VAR_GLOBAL   (* controller tags *)
   ACTIVE_MODE : ALIAS FOR N54[208].3;
   AFI : ALIAS FOR B3[7].15;
   AFITC : ALIAS FOR B3[15].15;
   AMAX_LEHR_SPD : ALIAS FOR I[81];
   APC_HOST_PERM : ALIAS FOR B3[0].7;
   AUX_xInitialize : BOOL;
   Axies : MOTION_GROUP; {access Read Only}
   B106 : DINT[1];
   B151 : DINT[20] := ([0] := 2#1111_1111_1111_1111_1111_1111_1111_1111, [1] := 2#1111_1111_1111_1111_1111_1111_1111_1111, [2] := 2#0000_0000_0000_0000_1111_1111_1111_1111);
        [0]   // Cross-break Zone 1 Bit shift file * INSIDE LEHR *
   B152 : DINT[50];
        [0]   // Cross-break Zone 2 Bit shift file ** LEHR EXIT **
        [8].14   // Crossbreak Zone 3 Crossbreak Active NEW Start bit
        [11].14   // Crossbreak Zone 3 Crossbreak Active OLD Start bit
   B153 : DINT[20] := ([0] := 2#1111_1111_1111_1111_1111_1111_1111_1111, [1] := 2#1111_1111_1111_1111_1111_1111_1111_1111, [2] := 2#1111_1111_1111_1111_1111_1111_1111_1111, [3] := 2#0000_0000_0000_0000_1111_1111_1111_1111);
        [0]   // Cross-break Zone 3 Bit shift file ** WASHER **
   B154 : DINT[20];
        [0]   // Cross-break Zone 4 Bit shift file * IMAGE AUTO *
        [1]   // Crossbreak
        [8].0   // Cross-break Zone 4 Bit shift file **
        [8].11   // Cross-break Zone 4 Bit shift file **
   B155 : DINT[20] := ([0] := 2#1111_1111_1111_1111_1111_1111_1111_1111, [1] := 2#1111_1111_1111_1111_1111_1111_1111_1111, [2] := 2#1111_1111_1111_1111_1111_1111_1111_1111, [3] := 2#1111_1111_1111_1111_1111_1111_1111_1111, [4] := 2#1111_1111_1111_1111_1111_1111_1111_1111, [5] := 2#1111_1111_1111_1111_1111_1111_1111_1111, [6] := 2#1111_1111_1111_1111_1111_1111_1111_1111, [7] := 2#1111_1111_1111_1111_1111_1111_1111_1111, [8] := 2#0000_0000_0000_0000_1111_1111_1111_1111);
        [0]   // Cross-break Zone 5 Bit shift file ** MAN. INSP **
        [1]   // Cross-break Zone 5 Bit shift file ** MAN. INSP **
        [1].11   // Cross-break Zone 5 Bit shift file APC Roll #1
        [4]   // Cross-break Zone 5 Bit shift file ** MAN. INSP **
        [4].0   // Cross-break Zone 5 Bit shift file APC Roll #2
        [5]   // Cross-break Zone 5 Bit shift file ** MAN. INSP **
   B175 : DINT[1];
   B176 : DINT[1] := ([0] := 2#0000_0000_0000_0000_0000_1100_0000_0000);
   B180 : DINT[10] := ([0] := 2#0000_0000_0000_0000_0000_1111_1000_0000, [1] := 2#0000_0000_0000_0000_0000_0000_0100_0000, [2] := 2#0000_0000_0000_0000_0000_0000_1000_0000, [4] := 2#0000_0000_0000_0000_0001_0000_0000_0000, [5] := 2#0000_0000_0000_0000_0000_0000_0011_0000);
   B3 : DINT[102] := ([0] := 2#0000_0000_0000_0000_0001_1001_0100_0000, [2] := 2#0000_0000_0000_0000_0000_0000_0000_0110, [7] := 2#0000_0000_0000_0000_0000_0000_0000_0001, [8] := 2#0000_0000_0000_0000_1100_0000_0000_0001, [10] := 2#0000_0000_0000_0000_0100_0000_0010_0001);
        [0].0   // Valid Flaw Data to Process
        [0].1   // Reversed Scanner
        [0].2   // Gun Number is Odd
        [0].3   // Cap Data Request ONS
        [0].4   // Reject (Flaw) PB ONS
        [0].5   // Gun Test Requested
        [0].7   // APC MACHINE Permissive to Run from Host
        [0].9   // HOST TRACKING Permissive to Operate lucor MSM machine
        [0].11   // Bridge in Down Position
        [0].12   // Bridge in Up Position
        [0].13   // Auto Down After Cross-Brk
        [0].14   // one shot
        [1].0   // one shot
        [1].1   // MARKING BRIDGE In final decel during downward travel
        [1].2   // No. 1 Crusher Chip Blower Manual Permissive
        [1].3   // No. 1 Crusher Chip Blower Automatic Permissive
        [1].12   // Cullet System M47B Fwd Direction Selected
        [1].13   // Cullet System M47B Rev Direction Selected
        [1].14   // Cullet System M37B Fwd Direction Selected
        [1].15   // Cullet Sytem M37B Rev Direction Selected
        [2].0   // One Shot
        [2].1   // ONE SHOT
        [2].2   // SPONGE ROLL MANUALLY ON
        [3].0   // Reliance Drive System Fault Permissive
        [3].1   // Cullet System Fault Permissive
        [4].0   // CROSS BREAK Present At Sub-surface Cutters
        [5].0   // temp debug for 1 m sync pulse
        [5].1   // temp debug for 1 m sync pulse
        [5].2   // LEHR SPEED Debug One shot
        [6].0   // One Shot for Accumulation of 20 50mm Pulses
        [6].1   // One Shot to Resume Accumulation of 50mm Pulses
        [7].0   // Crossbreak Active In Zones 1 or 2 Enable Beacons and Horn Lehr wall
        [7].15   // Always False
        [8].0   // Crossbreak 1 (Lehr) Fault Count One Shot
        [8].14   // North Chilled Water Blower Is Not On
        [8].15   // South Chilled Water Blower Is Not On
        [10].0   // APC Crossbreak or Estop Acknowledge to Reset Roller #1
        [10].1   // APC Early Crossbreak Drip Valve Shutoff
        [10].2   // LEHR SPEED one shot!
        [10].3   // LEHR SPEED one shot!
        [10].4   // Reliance Drive & Cullet System Alarm Horn Relay (Capping Rm)
        [10].5   // APC Crossbreak or Estop Acknowledge to Reset Roller #2
        [10].10   // APC Supply Flow Is Low Alarm
        [10].14   // Tony's Washer Disable Toggle Bit
        [10].15   // Always False
        [15].15   // Always false Tony Bit
        [80].0   // CT Lehr Conv have all stoped
        [0].6   // OK to Run Lehr AUX Conveyors
   B49 : DINT[100];
   B52 : DINT[100] := ([0] := 2#0000_0000_0000_0000_0000_0000_0000_0001);
        [0].0   // All of CT DRIVES Enable
   B73 : DINT[1];
        [0].1   // Two inch Tracking pulse For Lehr Speed
        [0].2   // Two inch Tracking pulse For trim Speed
   BIN_1B_EAST : ALIAS FOR O[112].12;
   BLOWER_ON : ALIAS FOR O[67].13;
   BOOTH_LIGHTS : ALIAS FOR N46[4];
   BRDG_EOT_LS_HI : ALIAS FOR I[12].3;
   BRDG_SLO_LS_HI : ALIAS FOR I[12].0;
   BRDG_SLO_LS_LO : ALIAS FOR I[12].1;
   BRIDGE_DOWN : ALIAS FOR B3[0].11;
   BRIDGE_DRV_FLT : ALIAS FOR I[17].0;
   BRIDGE_FIN_DEC : ALIAS FOR B3[1].1;
   BRIDGE_LO_LAMP : ALIAS FOR O[22].3;
   BRIDGE_MAN_INSP : ALIAS FOR I[18].4;
   BRIDGE_UP : ALIAS FOR B3[0].12;
   BRSH1_DN_FLT : ALIAS FOR I[43].1;
   BRSH1_DN_FWD : ALIAS FOR O[45].1;
   BRSH1_DN_REV : ALIAS FOR O[45].9;
   BRSH1_DN_SS1 : ALIAS FOR O[46].1;
   BRSH1_DN_SS2 : ALIAS FOR O[46].9;
   BRSH1_UP_FLT : ALIAS FOR I[43].0;
   BRSH1_UP_FWD : ALIAS FOR O[45].0;
   BRSH1_UP_REV : ALIAS FOR O[45].8;
   BRSH1_UP_SS1 : ALIAS FOR O[46].0;
   BRSH1_UP_SS2 : ALIAS FOR O[46].8;
   BRSH2_DN_FLT : ALIAS FOR I[43].3;
   BRSH2_DN_FWD : ALIAS FOR O[45].3;
   BRSH2_DN_REV : ALIAS FOR O[45].11;
   BRSH2_DN_SS1 : ALIAS FOR O[46].3;
   BRSH2_DN_SS2 : ALIAS FOR O[46].11;
   BRSH2_UP_FLT : ALIAS FOR I[43].2;
   BRSH2_UP_FWD : ALIAS FOR O[45].2;
   BRSH2_UP_REV : ALIAS FOR O[45].10;
   BRSH2_UP_SS1 : ALIAS FOR O[46].2;
   BRSH2_UP_SS2 : ALIAS FOR O[46].10;
   BT181_000 : MESSAGE;
        MessageParameters(ServiceCode := 16#004c, LocalElement := N125[0], ...)
   BT181_001 : MESSAGE;
        MessageParameters(ServiceCode := 16#004c, LocalElement := N125[62], ...)
   BT181_002 : MESSAGE;
        MessageParameters(ServiceCode := 16#004c, LocalElement := N125[123], ...)
   BT181_003 : MESSAGE;
        MessageParameters(ServiceCode := 16#004c, LocalElement := N125[183], ...)
   BT181_004 : MESSAGE;
        MessageParameters(ServiceCode := 16#004b, LocalElement := N124[0], ...)
   BT181_005 : MESSAGE;
        MessageParameters(ServiceCode := 16#004b, LocalElement := N124[62], ...)
   BT181_006 : MESSAGE;
        MessageParameters(ServiceCode := 16#004b, LocalElement := N124[123], ...)
   BT181_007 : MESSAGE;
        MessageParameters(ServiceCode := 16#004b, LocalElement := N124[183], ...)
   BT181_008 : MESSAGE;
        MessageParameters(ServiceCode := 16#004b, LocalElement := N124[250], ...)
   BT181_009 : MESSAGE;
        MessageParameters(ServiceCode := 16#004c, LocalElement := N125[350], ...)
   BT181_010 : MESSAGE;
        MessageParameters(ServiceCode := 16#004b, LocalElement := N124[350], ...)
   BT181_011 : MESSAGE;
   BT181_012 : MESSAGE;
        MessageParameters(LocalElement := N15[60], ...)
   BT181_013 : MESSAGE;   // MB TO M2 BT of MMI Data To New CLX PLC
        MessageParameters(LocalElement := N7[180], ...)
   BT181_014 : MESSAGE;   // M2 TO MB BT of MMI Data from New CLX PLC
        MessageParameters(LocalElement := N7[160], ...)
   BT41_000 : MESSAGE;   // VHSC BTR
        .EN   // VHSC BTR Enabled
        MessageParameters(ServiceCode := 16#004b, LocalElement := N42[71], ...)
   BT41_001 : MESSAGE;   // VHSC BTW
        .EN   // VHSC BTW Enabled
        MessageParameters(ServiceCode := 16#004c, LocalElement := N42[1], ...)
   BT41_002 : MESSAGE;
        MessageParameters(LocalElement := N45[21], ...)
   BT41_003 : MESSAGE;
        MessageParameters(LocalElement := N45[1], ...)
   BT41_004 : MESSAGE;
   BT41_005 : MESSAGE;
   BT41_006 : MESSAGE;   // Block Transfer Read Control for Analog Input Card in Washer Panel
        MessageParameters(ServiceCode := 16#004b, LocalElement := N61[1], ...)
   BT41_007 : MESSAGE;   // Block Transfer Write Control for Analog Input Card in Washer Panel
        MessageParameters(ServiceCode := 16#004c, LocalElement := N61[51], ...)
   C183 : COUNTER[3] := ([0].PRE := 1, [0].CU := 1, [1].PRE := 7, [1].CU := 1, [2].PRE := 3, [2].CU := 1);
   C1_ACK : ALIAS FOR N54[260].14;
   C1_ACTIVE_LAMP : ALIAS FOR N54[260].0;
   C1_BEACON : ALIAS FOR O[27].6;
   C1_BEACON2 : ALIAS FOR O[47].10;
   C1_HORN : ALIAS FOR O[27].5;
   C1_NTH_IN_LMP : ALIAS FOR N54[260].10;
   C1_NTH_IN_PE : ALIAS FOR N54[260].6;
   C1_NTH_IN_SS : ALIAS FOR N54[260].2;
   C1_NTH_OUT_LMP : ALIAS FOR N54[260].9;
   C1_NTH_OUT_PE : ALIAS FOR N54[260].5;
   C1_NTH_OUT_SS : ALIAS FOR N54[260].1;
   C1_PNL_FLT : ALIAS FOR I[113].2;
   C1_STH_IN_LMP : ALIAS FOR N54[260].12;
   C1_STH_IN_PE : ALIAS FOR N54[260].8;
   C1_STH_IN_SS : ALIAS FOR N54[260].4;
   C1_STH_OUT_LMP : ALIAS FOR N54[260].11;
   C1_STH_OUT_PE : ALIAS FOR N54[260].7;
   C1_STH_OUT_SS : ALIAS FOR N54[260].3;
   C253 : COUNTER[100];
   C2_ACTIVE_LAMP : ALIAS FOR N54[261].0;
   C2_NTH_IN_LMP : ALIAS FOR N54[261].10;
   C2_NTH_IN_PE : ALIAS FOR N54[261].6;
   C2_NTH_IN_SS : ALIAS FOR N54[261].2;
   C2_NTH_OUT_LMP : ALIAS FOR N54[261].9;
   C2_NTH_OUT_PE : ALIAS FOR N54[261].5;
   C2_NTH_OUT_SS : ALIAS FOR N54[261].1;
   C2_PNL_FLT : ALIAS FOR I[113].3;
   C2_STH_IN_LMP : ALIAS FOR N54[261].12;
   C2_STH_IN_PE : ALIAS FOR N54[261].8;
   C2_STH_IN_SS : ALIAS FOR N54[261].4;
   C2_STH_OUT_LMP : ALIAS FOR N54[261].11;
   C2_STH_OUT_PE : ALIAS FOR N54[261].7;
   C2_STH_OUT_SS : ALIAS FOR N54[261].3;
   C3_ACTIVE_LAMP : ALIAS FOR N54[262].0;
   C3_NTH_IN_LMP : ALIAS FOR N54[262].10;
   C3_NTH_IN_PE : ALIAS FOR N54[262].6;
   C3_NTH_IN_SS : ALIAS FOR N54[262].2;
   C3_NTH_OUT_LMP : ALIAS FOR N54[262].9;
   C3_NTH_OUT_PE : ALIAS FOR N54[262].5;
   C3_NTH_OUT_SS : ALIAS FOR N54[262].1;
   C3_PNL_FLT : ALIAS FOR I[113].4;
   C3_STH_IN_LMP : ALIAS FOR N54[262].12;
   C3_STH_IN_PE : ALIAS FOR N54[262].8;
   C3_STH_IN_SS : ALIAS FOR N54[262].4;
   C3_STH_OUT_LMP : ALIAS FOR N54[262].11;
   C3_STH_OUT_PE : ALIAS FOR N54[262].7;
   C3_STH_OUT_SS : ALIAS FOR N54[262].3;
   C3_STP : ALIAS FOR O[35].10;
   C4_NTH_IN_PE : ALIAS FOR N54[263].6;
   C4_NTH_IN_SS : ALIAS FOR N54[263].2;
   C4_NTH_OUT_PE : ALIAS FOR N54[263].5;
   C4_NTH_OUT_SS : ALIAS FOR N54[263].1;
   C4_PNL_FLT : ALIAS FOR I[113].1;
   C4_STH_IN_PE : ALIAS FOR N54[263].8;
   C4_STH_OUT_PE : ALIAS FOR N54[263].7;
   C5 : COUNTER[100] := ([0].PRE := 200, [1].PRE := 2, [2].PRE := 52, [2].ACC := 29, [3].PRE := 30000, [3].ACC := 2, [4].PRE := 30000, [5].PRE := 30000, [6].PRE := 1000, [6].ACC := 423, [7].PRE := 30000, [8].PRE := 1000, [8].ACC := 112, [8].CU := 1, [10].PRE := 30000, [12].PRE := 30000, [13].PRE := 32767, [13].ACC := 1912, [14].ACC := 74, [14].DN := 1, [15].ACC := 54, [15].DN := 1, [16].ACC := 33, [16].DN := 1, [17].ACC := 27, [17].DN := 1, [20].PRE := 1000, [20].ACC := 1748, [20].DN := 1, [21].PRE := 1000, [21].ACC := 13747, [21].DN := 1, [21].OV := 1, [25].PRE := 1000, [25].ACC := 853, [26].PRE := 10000, [26].ACC := 3, [27].PRE := 10000, [27].ACC := 4, [27].CU := 1, [28].PRE := 10000, [28].ACC := 4, [28].CU := 1, [29].PRE := 10000, [29].ACC := 4, [29].CU := 1, [30].PRE := 10000, [30].ACC := 4, [30].CU := 1, [31].PRE := 10000, [31].ACC := 2145, [32].PRE := 10000, [32].ACC := 4, [32].CU := 1, [33].PRE := 10000, [34].PRE := 10000, [34].ACC := 4, [35].PRE := 10000, [35].ACC := 2786, [36].PRE := 10000,
        [36].ACC := 4, [37].PRE := 10000, [37].ACC := 2743, [38].PRE := 10000, [38].ACC := 4, [39].PRE := 10000, [39].ACC := 2790, [40].PRE := 10000, [40].ACC := 4, [41].PRE := 10000, [41].ACC := 2693, [42].PRE := 10000, [42].ACC := 4, [43].PRE := 10000, [43].ACC := 5802, [44].PRE := 10000, [44].ACC := 4, [45].PRE := 10000, [45].ACC := 11749, [45].DN := 1, [46].PRE := 10000, [46].ACC := 4, [46].DN := 1, [46].OV := 1, [47].PRE := 10000, [47].ACC := 478, [48].PRE := 10000, [48].ACC := 4, [49].PRE := 10000, [49].ACC := 6623, [50].PRE := 10000, [50].ACC := 4424, [51].PRE := 10000, [51].ACC := 734, [52].PRE := 10000, [52].ACC := 5426, [53].PRE := 10000, [53].ACC := 783, [54].PRE := 10000, [54].ACC := 3735, [55].PRE := 10000, [55].ACC := 733, [56].PRE := 10000, [56].ACC := 3661, [57].PRE := 10000, [57].ACC := 727, [58].PRE := 1000, [58].ACC := 251, [58].CU := 1, [70].PRE := 10000, [70].CU := 1, [71].PRE := 10000, [71].ACC := 4, [71].CU := 1, [72].PRE := 10000, [72].CU := 1, [73].PRE := 10000, [73].ACC := 4, [73].CU := 1, [74].PRE := 10000,
        [74].CU := 1, [75].PRE := 10000, [75].ACC := 4, [75].CU := 1, [76].PRE := 10000, [76].CU := 1, [77].PRE := 10000, [77].ACC := 4, [77].CU := 1, [78].PRE := 1000, [78].ACC := 607, [79].PRE := 1000, [79].ACC := 300, [80].PRE := 1000, [80].ACC := 337, [81].PRE := 1000, [81].ACC := 1033, [81].DN := 1, [82].PRE := 1000, [82].ACC := 146, [83].PRE := 1000, [83].ACC := 63, [84].PRE := 1000, [84].ACC := 2159, [84].DN := 1, [85].PRE := 1000, [85].ACC := 553, [90].PRE := 10000, [90].ACC := 8, [91].PRE := 10000, [93].PRE := 1000, [93].ACC := 338, [93].CU := 1, [94].PRE := 100, [95].PRE := 100, [96].PRE := 100, [96].ACC := 65, [97].PRE := 100, [97].ACC := 65, [98].PRE := 10000, [98].ACC := 6222, [99].PRE := 1000, [99].ACC := 520, [99].CU := 1);
        [6]   // TEMP Counter for Number of Times South OUT Sensor gets Disabled
        [13]   // Reliance Drive & Cullet System Alarm Horn (Capping) Conter
        [20]   // DEBUG: Number Of Times Capping Lehr Speed is Greater than Automax Speed plus 15IPM
        [21]   // TEMP DEBUG NUMBER OF TIMES 1M SYNC PULSE PERIOD IS LESS THAN 8 SEC
        [25]   // M2-->>MB Counts number of Times Mainline Backup to Trim Deck Occurs
        [26]   // CB Zone 1 (Lehr) North Outside Debounce Counter
        [27]   // CB Zone 1 (Lehr) North Outside Fault Counter
        [28]   // CB Zone 1 (Lehr) North Inside Debounce Counter
        [29]   // CB Zone 1 (Lehr) North Inside Fault Counter
        [30]   // CB Zone 1 (Lehr) South Outside Debounce Counter
        [31]   // CB Zone 1 (Lehr) South Outside Fault Counter
        [32]   // CB Zone 1 (Lehr) South Inside Debounce Counter
        [33]   // CB Zone 1 (Lehr) South Inside Fault Counter
        [34]   // CB Zone 2 (Crusher 1) North Outside Debounce Counter
        [35]   // CB Zone 2 (Crusher 1) North Outside Fault Counter
        [36]   // CB Zone 2 (Crusher 1) North Inside Debounce Counter
        [37]   // CB Zone 2 (Crusher 1) North Inside Fault Counter
        [38]   // CB Zone 2 (Crusher 1) South Outside Debounce Counter
        [39]   // CB Zone 2 (Crusher 1) South Outside Fault Counter
        [40]   // CB Zone 2 (Crusher 1) South Inside Debounce Counter
        [41]   // CB Zone 2 (Crusher 1) South Inside Fault Counter
        [42]   // CB Zone 3 (washer) North Outside Debounce Counter
        [43]   // CB Zone 3 (washer) North Outside Fault Counter
        [44]   // CB Zone 3 (washer) North Inside Debounce Counter
        [45]   // CB Zone 3 (washer) North Inside Fault Counter
        [45].ACC   // Z2 NO
        [46]   // CB Zone 3 (washer) South Outside Debounce Counter
        [46].ACC   // Z2 NI
        [47]   // CB Zone 3 (washer) South Outside Fault Counter
        [47].ACC   // Z2 SO
        [48]   // CB Zone 3 (washer) South Inside Debounce Counter
        [48].ACC   // Z2 SI
        [49]   // CB Zone 3 (washer) South Inside Fault Counter
        [50].ACC   // Z3 NO
        [51]   // CB Zone 4 (Inspection Booth) North Outside Fault Counter
        [51].ACC   // Z3 NI
        [52].ACC   // Z3 SO
        [53]   // CB Zone 4 (Inspection Booth) North Inside Fault Counter
        [53].ACC   // Z3 NI
        [54].ACC   // Z4 SI
        [55]   // CB Zone 4 (Inspection Booth) South Outside Fault Counter
        [55].ACC   // Z4 SO
        [56].ACC   // Z4 NI
        [57]   // CB Zone 4 (Inspection Booth) South Inside Fault Counter
        [57].ACC   // Z4 NO
        [71].ACC   // Z5 NO
        [73].ACC   // Z5 SI
        [75].ACC   // Z5 SO
        [77].ACC   // Z5 SI
        [90]   // Temporary Counter to Monitor CT Master Drive Fault Contact 0 ON 03/11/08
        [94]   // I/O STATUS FILE: Rack 12 Group 6 FAULT
        [95]   // I/O STATUS FILE: Rack 12 Group 4 FAULT
        [96]   // I/O STATUS FILE: Rack 12 Group 2 FAULT
        [97]   // I/O STATUS FILE: Rack 12 Group 0 FAULT
        [98]   // Glass Travel Pulse Count (Counts 50mm Pulses reset @ 10000)
        [99]   // BRUSH 1 DRIVE FAULTS
   C5_ACTIVE_LAMP : ALIAS FOR N54[264].0;
   C5_MARKING_CB : ALIAS FOR N54[264].15;
   C5_NTH_IN_LMP : ALIAS FOR N54[264].10;
   C5_NTH_IN_PE : ALIAS FOR N54[264].6;
   C5_NTH_IN_SS : ALIAS FOR N54[264].2;
   C5_NTH_OUT_LMP : ALIAS FOR N54[264].9;
   C5_NTH_OUT_PE : ALIAS FOR N54[264].5;
   C5_NTH_OUT_SS : ALIAS FOR N54[264].1;
   C5_STH_IN_LMP : ALIAS FOR N54[264].12;
   C5_STH_IN_PE : ALIAS FOR N54[264].8;
   C5_STH_IN_SS : ALIAS FOR N54[264].4;
   C5_STH_OUT_LMP : ALIAS FOR N54[264].11;
   C5_STH_OUT_PE : ALIAS FOR N54[264].7;
   C5_STH_OUT_SS : ALIAS FOR N54[264].3;
   CAP_AHR_TMR : ALIAS FOR T4[6];
   CAP_ALM_HORN : ALIAS FOR O[11].2;
   CAW_OK_BIT_W_PLC : ALIAS FOR N251[901].0;
   CAWSV_ON_BIT_TO_WPLC : ALIAS FOR N251[900].0;
   CB_AT_SS_CUTTERS : ALIAS FOR B3[4].0;
   CBF_START_B : ALIAS FOR I[65].5;
   CBF_START_T : ALIAS FOR I[65].4;
   CBF_STOP_B : ALIAS FOR I[65].7;
   CBF_STOP_T : ALIAS FOR I[65].6;
   CHIP_BLOW_A : ALIAS FOR B3[1].3;
   CHIP_BLOW_M : ALIAS FOR B3[1].2;
   CHIP_BLOW_TMR : ALIAS FOR T51[9];
   CNV10_PROCST : ALIAS FOR I[19].9;
   CNV11_PROCST : ALIAS FOR I[3].1;
   CNV12_PROCST : ALIAS FOR I[3].2;
   CNV13_PROCST : ALIAS FOR I[3].3;
   CNV14_PROCST : ALIAS FOR I[3].4;
   CNV15_PROCST : ALIAS FOR I[3].5;
   CNV16_PROCST : ALIAS FOR I[3].7;
   CNV17_PROCST : ALIAS FOR I[3].8;
   CNV1_PROCST : ALIAS FOR I[19].0;
   CNV2_PROCST : ALIAS FOR I[19].1;
   CNV3_PROCST : ALIAS FOR I[19].2;
   CNV4_PROCST : ALIAS FOR I[19].3;
   CNV5_PROCST : ALIAS FOR I[19].4;
   CNV6_PROCST : ALIAS FOR I[19].5;
   CNV7_PROCST : ALIAS FOR I[19].6;
   CNV8_PROCST : ALIAS FOR I[19].7;
   CNV9_PROCST : ALIAS FOR I[19].8;
   ConsumedFromCullet : UDT_CONSUMED_CULLET;
   ConsumedFromMCC1300 : UDT_CONSUMED_NEXT := (iM2toMB_2 := 132, iM2toMB_4 := 2048);
   CPU_FaultRecord : SYS_FaultRecord;
   CPU_LastFaultRecord : SYS_FaultRecord;
   CR1_0FF_LAMP : ALIAS FOR O[67].9;
   CR1_ALM : ALIAS FOR I[65].1;
   CR1_AUTO : ALIAS FOR I[64].13;
   CR1_AUTO_MODE : ALIAS FOR N54[240].1;
   CR1_CONT_FAIL : ALIAS FOR N54[240].4;
   CR1_CULLET_FAIL : ALIAS FOR N54[240].6;
   CR1_DNET_SS1 : ALIAS FOR N179[18];
   CR1_DNET_SS2 : ALIAS FOR N179[30];
   CR1_DOWN_PROX : ALIAS FOR I[64].11;
   CR1_DOWN_PWRLOS : ALIAS FOR N54[240].10;
   CR1_DOWN_RLY : ALIAS FOR O[67].1;
   CR1_DROP_COND : ALIAS FOR N54[240].13;
   CR1_DRV_FLT_LMP : ALIAS FOR O[66].8;
   CR1_DRV_FLT_RLY : ALIAS FOR O[66].9;
   CR1_DWN_PROX : ALIAS FOR N54[240].14;
   CR1_ESTOP : ALIAS FOR N54[240].3;
   CR1_FLT : ALIAS FOR I[65].0;
   CR1_FRSTSCN_TMR : ALIAS FOR T51[11];
   CR1_FWD : ALIAS FOR O[66].0;
   CR1_MAN_LOWER : ALIAS FOR I[64].15;
   CR1_MAN_MODE : ALIAS FOR N54[240].2;
   CR1_MAN_RAISE : ALIAS FOR I[64].14;
   CR1_NODROP_COND : ALIAS FOR N54[240].0;
   CR1_ON_LAMP : ALIAS FOR O[67].8;
   CR1_RUN_ENABLE : ALIAS FOR O[117].4;
   CR1_SS1 : ALIAS FOR O[66].2;
   CR1_SS2 : ALIAS FOR O[66].4;
   CR1_SS3 : ALIAS FOR O[66].6;
   CR1_START_PB : ALIAS FOR I[65].12;
   CR1_STOP_PB : ALIAS FOR I[65].13;
   CR1_TEST_PB : ALIAS FOR I[65].3;
   CR1_UP_PROX : ALIAS FOR I[64].12;
   CR1_UP_RLY : ALIAS FOR O[67].0;
   CR1_UPT_PROX : ALIAS FOR N54[240].15;
   CULL_FLT : ALIAS FOR B3[3].1;
   CULLET_FLT_PL : ALIAS FOR O[11].1;
   CURR_LSD : ALIAS FOR N42[74];
   CURR_MSD : ALIAS FOR N42[73];
   CURR_SYNC : ALIAS FOR N7[2];
   DateTime : DINT[7] := ([0] := 2023, [1] := 6, [2] := 9, [3] := 15, [4] := 17, [5] := 5, [6] := 737882);   // DINT array tag for retrieve wallclock time through GSV created during conversion
        [0]   // Year
        [1]   // Month
        [2]   // Day
        [3]   // Hour
        [4]   // Minute
        [5]   // Second
        [6]   // Microsecond
   DISABLE_REL : ALIAS FOR N46[3];
   DISTANCE : ALIAS FOR N7[1];
   DIV_POSITION : ALIAS FOR I[24].12;
   DIVERTER_POS1 : ALIAS FOR O[116].8;
   DRIVE_FAULT_PRESENT : BOOL; {access Read Only}
   ECLIPSE_OFF : ALIAS FOR N54[208].2;
   ECLIPSE_ON : ALIAS FOR N54[208].1;
   EMERGENCY_OK : BOOL;
   F58 : REAL[20] := ([0] := 5063.717);
        [0]   // APC Calculated Freq for APC Roller [Hz * 100]
   F74 : REAL[2] := ([0] := 13.333333, [1] := 0.15);
   F8 : REAL[20] := ([5] := 3.125);
        [5]   // SHEET TEMPERATURE: Tuning Factor to adjust PLC Value to match LED Display Unit
   F96 : REAL[50] := ([0] := 268.34647, [1] := 268.34647, [5] := 118.346466, [6] := 418.34647, [9] := 270.6, [10] := 270.6, [11] := 268.34647, [12] := 1.94725, [14] := 285.6, [20] := 268.34647, [21] := 268.34647, [22] := 268.34647, [23] := 268.34647, [24] := 268.34647, [25] := 268.34647, [26] := 268.34647, [27] := 268.34647, [28] := 268.34647, [29] := 268.34647, [30] := 270.6, [40] := 268.34647, [41] := 268.34647, [42] := 268.34647, [43] := 268.34647, [44] := 268.34647, [45] := 268.34647, [46] := 268.34647, [47] := 268.34647, [48] := 268.34647, [49] := 268.34647);
        [0]   // LEHR SPEED Current lehr Speed used Setting Speed of drives
        [1]   // LEHR SPEED Average lehr Speed Calculated from Sample table
        [5]   // LEHR SPEED Current Lehr Lower Limit
        [6]   // LEHR SPEED Current Lehr Speed upper Limit
        [9]   // LEHR SPEED Last lehr Speed Reset value
        [10]   // LEHR SPEED Information Received from Reliance AutoMax
        [11]   // LEHR SPEED Information Received from Reliance Capping system
        [14]   // DEBUG USAGE Lehr Speed from Automax Plus 15 IPM
        [20]   // LEHR SPEED Table of Speed samples Over last ten Seconds
        [21]   // LEHR SPEED Table of Lehr speed Samples over Ten seconds
   FAST_FLASH : ALIAS FOR T51[2];
   FFLASH_SLAVE : ALIAS FOR T51[3];
   FIRST_SCAN : ALIAS FOR S[1].15;
   FLAW_HEAD : ALIAS FOR N43[200];
   FLAW_LANE : ALIAS FOR N43[201];
   FLAW_OFF : ALIAS FOR N43[202];
   FLAW_OUT : ALIAS FOR N7[5];
   FLAW_POS : ALIAS FOR N7[4];
   FLAW_QUEUE : ALIAS FOR N7[9];
   FLAW_XLAT : ALIAS FOR N7[6];
   FLOW_CLK_LSD : ALIAS FOR N7[10];
   FLOW_CLK_MSD : ALIAS FOR N7[11];
   ForceStatus : INT;   // INT tag to retrieve Force enabled value through GSV created during conversion
   From_Cullet : DINT[10];
   GENERATOR_ON : ALIAS FOR N54[240].11;
   GENERATOR_RUN : ALIAS FOR I[65].15;
   GOOD_FLAW : ALIAS FOR B3[0].0;
   GP_M225_AccessArea : GP_AccessArea := (IN_xConditionOkAccess := 1); {access None}
   GP_M225_AccessArea_STC : GP_AccessArea_STC := (OSR_xRemoveAccess := 1, OSR_xRemoveAccessNotAccepted := 1, tmON_ForceAccess.PRE := 5000); {access None}
   GP_NetDiag : GP_NetworkDiag;
   GP_OB_InitializeDiag : GP_OB_Initialize := (OUT_dExecutionTime_ms := 500, OUT_dMaxExecutionTime_ms := 1033885, OUT_xOs_100ms := 1, OUT_xOs_200ms := 1, OUT_xOs_400ms := 1, OUT_xOs_500ms := 1, OUT_xOs_800ms := 1, OUT_xClock_100ms := 1, OUT_xClock_200ms := 1, OUT_xClock_400ms := 1, OUT_xClock_500ms := 1, OUT_xClock_800ms := 1, OUT_xClock_1s := 1, OUT_xClock_5s := 1, OUT_xClock_10s := 1, OUT_xClock_30s := 1, OUT_xClock_1h := 1, OUT_xDebugON := 1);
   GP_OB_InitializeDiag_STC : GP_OB_Initialize_STC := (dElapsed_1h_ms := 7496626, dElapsed_1min_ms := 56626, dElapsed_1s_ms := 626, dElapsed_2min_ms := 56626, dElapsed_2s_ms := 626, dElapsed_5s_ms := 1626, dElapsed_10min_ms := 296626, dElapsed_10s_ms := 6626, dElapsed_30min_ms := 296626, dElapsed_30s_ms := 26626, dElapsed_100ms_ms := 75523026, dElapsed_200ms_ms := 57149426, dElapsed_400ms_ms := 20402226, dElapsed_500ms_ms := 2028626, dElapsed_800ms_ms := 626, dlLastExecValue_us := 499964, rReminder_ms := -0.35214233, lwOldStartTime[0] := -592654905, lwOldStartTime[1] := 392627, lwStartTime[0] := -592654905, lwStartTime[1] := 392627);
   GP_OB_InitializeMain : GP_OB_Initialize := (OUT_dExecutionTime_ms := 10, OUT_dMaxExecutionTime_ms := 11, OUT_xOs_100ms := 1, OUT_xOs_200ms := 1, OUT_xClock_200ms := 1, OUT_xClock_800ms := 1, OUT_xClock_1s := 1, OUT_xClock_2s := 1, OUT_xClock_5s := 1, OUT_xClock_10s := 1, OUT_xClock_30s := 1, OUT_xClock_2min := 1, OUT_xClock_10min := 1, OUT_xDebugON := 1);
   GP_OB_InitializeMain_STC : GP_OB_Initialize_STC := (dElapsed_1h_ms := 4478668, dElapsed_1min_ms := 38668, dElapsed_1s_ms := 668, dElapsed_2min_ms := 38668, dElapsed_2s_ms := 668, dElapsed_5s_ms := 3668, dElapsed_10min_ms := 278668, dElapsed_10s_ms := 8668, dElapsed_30min_ms := 878668, dElapsed_30s_ms := 8668, dElapsed_100ms_ms := 68, dElapsed_200ms_ms := 68, dElapsed_400ms_ms := 268, dElapsed_500ms_ms := 168, dElapsed_800ms_ms := 268, dlLastExecValue_us := 9789, rReminder_ms := -0.0073947906, lwOldStartTime[0] := -593976054, lwOldStartTime[1] := 392627, lwStartTime[0] := -593976054, lwStartTime[1] := 392627);
   GUN_INDEX : ALIAS FOR N7[0];
   HMI_Alarm_Presence : BOOL;   // HMI_Alarm_Presence
   HMI_Alarm_Reset : BOOL;   // HMI_Alarm_Reset
   HMI_Alarms_0 : BOOL[32];   // HMI Alarms
   HMI_Alarms_1 : BOOL[32];   // HMI Alarms
   HMI_Alarms_2 : BOOL[32];   // HMI Alarms
   HMI_Alarms_3 : BOOL[32];   // HMI Alarms
   HMI_Alarms_4 : BOOL[32];   // HMI Alarms
   HMI_Alarms_5 : BOOL[32];   // HMI Alarms
   HMI_Alarms_6 : BOOL[32];   // HMI Alarms
   HMI_Alarms_7 : BOOL[32];   // HMI Alarms
   HMI_Alarms_8 : BOOL[32];   // HMI Alarms
   HMI_Alarms_9 : BOOL[32];   // HMI Alarms
   HMI_Always_ON : BOOL := 1;   // HMI Always ON
   HMI_MAN_CMD_WR : UDT_MAN_CMD_WR; {access Read Only}
   HMI_MOTOR_HMR : UDT_MOTOR_HMR; {access Read Only}
   HOST_DATA_REQ : ALIAS FOR N43[209].0;
   HOST_IAL_ALARM : ALIAS FOR N43[209].6;
   HOST_IAL_WD : ALIAS FOR N43[209].7;
   HOST_NWDATA_TMR : ALIAS FOR T4[3];
   I : INT[128] := ([14] := 2#0000_0000_0010_0001, [15] := 2#0000_0000_0010_0001, [16] := 2#0000_0000_0000_0100, [17] := 2#1001_0000_0100_0000, [42] := 2#0000_0100_1110_1110, [43] := 2#0000_0000_1011_0000, [49] := 2#0000_0000_0010_0001, [65] := 2#1000_0001_1100_0001, [80] := 2#0011_0110_1111_0011, [81] := 2#0000_1010_1001_0010, [83] := 2#0000_0000_0001_1111, [121] := 2#0000_0000_1000_0100, [123] := 2#0000_1000_0000_0000);
        [42].9   // VMCC W1 Alarm Reset (NOT USED ANYMORE)
        [62].14   // SPARE
        [120]   // M2 --> MB
        [0].15   // PANEL C1 M47B Conv Forward Selector (INCLINE)
        [1].8   // PANEL C1 M47B Conv Reverse Selector (INCLINE)
        [3].0   // Transfer 1 Belt Process Stop Enabled
        [3].1   // Conveyor 11 Process Stop Enabled
        [3].2   // Conveyor 12 Process Stop Enabled
        [3].3   // Conveyor 13 Process Stop Enabled
        [3].4   // Conveyor 14 Process Stop Enabled
        [3].5   // Conveyor 15 Process Stop Enabled
        [3].6   // Transfer 1A Bel Process Stop Enabled
        [3].7   // Conveyor 16 Process Stop Enabled
        [3].8   // Conveyor 17 Process Stop Enabled
        [12].0   // Bridge Top Slow Down L.S.
        [12].1   // Bridge bottom Slow L.S.
        [12].3   // Bridge Top E.O.T. L.S.
        [12].14   // Reliance Data Request
        [12].15   // Reliance Two inch Lehr Pulse
        [16].0   // ISRA 5D 24VDC OK
        [16].4   // ISRA 5D 12V DC OK
        [16].5   // ISRA 5D System Ok
        [16].6   // ISRA 5D System Warning
        [16].7   // ISRA 5D System Error 1
        [16].8   // ISRA 5D System Error 2
        [16].9   // VMCC MB Alarm Silence
        [16].10   // VMCC MB Alarm Reset
        [16].14   // ISRA 5D System Crossbreak
        [17].1   // South Chilled Water Blower Off PB I02105
        [17].2   // North Subsurface Cutter Alarm Signal
        [17].3   // South Subsurface Cutter Alarm Signal
        [17].4   // South Chilled Water Blower On PB I02104
        [17].5   // South Chilled Water Blower Off PB I02105
        [17].7   // South Chilled Water Blower VFD is Running Without Faults
        [17].9   // Inspection in Manual Mode
        [17].10   // North Chilled Water Blower On PB I02112
        [17].11   // North Chilled Water Blower Off PB I02113
        [16].3   // ISRA 5D System Watchdog (NOT USED)
        [17].13   // North Chilled Water Blower VFD is Running Without Faults
        [17].14   // TO BE VALORIZED FROM MCC1200 Data Request From New Cutting System (Data Request from Reliance)
        [18].2   // SPARE (APC Reset Button After Crossbreak)
        [18].4   // SPARE (Inspection in Manual Mode)
        [16].1   // Spare
        [18].3   // SPARE (APC ON/OFF (0=OFF) (1=ON))
        [19].0   // Conveyor 1 Process Stop Enabled
        [19].1   // Conveyor 2 Process Stop Enabled
        [19].2   // Conveyor 3 Process Stop Enabled
        [19].3   // Conveyor 4 Process Stop Enabled
        [19].4   // Conveyor 5 Process Stop Enabled
        [19].5   // Conveyor 6 Process Stop Enabled
        [19].6   // Conveyor 7 Process Stop Enabled
        [19].7   // Conveyor 8 Process Stop Enabled
        [19].8   // Conveyor 9 Process Stop Enabled
        [19].9   // Conveyor 10 Process Stop Enabled
        [24].0   // CRSSBRK ZONE 1 North Outside Bypass Switch
        [24].1   // CRSSBRK ZONE 1 North Inside Bypass Switch
        [24].2   // CRSSBRK ZONE 1 South Outside Bypass Switch
        [24].3   // CRSSBRK ZONE 1 South Inside Bypass Switch
        [24].4   // CRSSBRK ZONE 1 North Outside Photo-cell
        [24].5   // CRSSBRK ZONE 1 North Inside Photo-cell
        [24].6   // CRSSBRK ZONE 1 South Outside Photo-cell
        [24].7   // CRSSBRK ZONE 1 South Inside Photo-cell
        [24].8   // Cullet System M37B Fwd Direction Selector (Outside)
        [24].9   // Cullet System M37B Rev Direction Selector (Outside)
        [24].10   // Cullet System M47B Fwd Direction Selector (Outside)
        [24].11   // Cullet System M47B Rev Direction Selector (Outside)
        [24].12   // Diverter Position Selector At Cullet Op Panel
        [26].0   // CRSSBRK ZONE 2 North Outside Bypass Switch
        [26].1   // CRSSBRK ZONE 2 North Inside Bypass Switch
        [26].2   // CRSSBRK ZONE 2 South Outside Bypass Switch
        [26].3   // CRSSBRK ZONE 2 South Inside Bypass Switch
        [26].4   // CRSSBRK ZONE 2 North Outside Photo-cell
        [26].5   // CRSSBRK ZONE 2 North Inside Photo-cell
        [26].6   // CRSSBRK ZONE 2 South Outside Photo-cell
        [26].7   // CRSSBRK ZONE 2 South Inside Photo-cell
        [28].0   // CRSSBRK ZONE 3 North Outside Bypass Switch
        [28].1   // CRSSBRK ZONE 3 North Inside Bypass Switch
        [28].2   // CRSSBRK ZONE 3 South Outside Bypass Switch
        [28].3   // CRSSBRK ZONE 3 South Inside Bypass Switch
        [28].4   // CRSSBRK ZONE 3 North Outside Photo-cell
        [28].5   // CRSSBRK ZONE 3 North Inside Photo-cell
        [28].6   // CRSSBRK ZONE 3 South Outside Photo-cell
        [28].7   // CRSSBRK ZONE 3 South Inside Photo-cell
        [30].13   // CRSSBRK ZONE 4 Adapter power ON
        [30].15   // CRSSBRK ZONE 4 Output power ON
        [30].12   // IMAGE AUTO Retro-cover Closed Prox
        [32].0   // CRSSBRK ZONE 5 North Outside Bypass Switch
        [32].1   // CRSSBRK ZONE 5 North Inside Bypass Switch
        [32].2   // CRSSBRK ZONE 5 South Outside Bypass Switch
        [32].3   // CRSSBRK ZONE 5 South Inside Bypass Switch
        [32].4   // CRSSBRK ZONE 5 North Outside Photo-cell
        [32].5   // CRSSBRK ZONE 5 North Inside Photo-cell
        [32].6   // CRSSBRK ZONE 5 South Outside Photo-cell
        [32].7   // CRSSBRK ZONE 5 South Inside Photo-cell
        [32].8   // APC #1 Reset Button After Crossbreak
        [32].9   // APC Spray system OFF (1=OFF) (0=ON)
        [32].10   // APC #2 Reset Button After Crossbreak changed 22Mar2019TC
        [32].11   // APC Spray System Supply Flow Low (From SMC flow meter)
        [34].0   // MANUAL INSPCTN Booth Flaw Push-Button
        [34].1   // MANUAL INSPCTN Booth Reject Push-Button
        [34].3   // LOW-E Inspection Catwalk: Spray Zone 1 Pushbutton
        [34].4   // LOW-E Inspection Catwalk: Spray Zone 2 Pushbutton
        [34].5   // LOW-E Inspection Catwalk: Spray Zone 3 Pushbutton
        [34].6   // LOW-E Inspection Catwalk: Spray Zone 4 Pushbutton
        [34].7   // LOW-E Inspection Catwalk: Spray Zone 5 Pushbutton
        [34].8   // LOW-E Inspection Catwalk: Pulse Entire Ribbon Pushbutton
        [58].12   // SPARE
        [58].13   // SPARE
        [58].10   // SPARE
        [58].15   // SPARE
        [60].15   // SPARE
        [58].9   // SPARE
        [56].15   // SPARE
        [58].11   // SPARE
        [58].14   // SPARE
        [43].0   // VMCC W1 Upper Brush #1 Drive fault
        [43].1   // VMCC W1 Lower Brush #1 Drive fault
        [43].2   // VMCC W1 Upper Brush #2 Drive fault
        [43].3   // VMCC W1 Lower Brush #2 Drive fault
        [43].6   // VMCC W1 SPARE
        [43].7   // VMCC W1 SPARE
        [43].8   // VMCC W1 SPARE
        [43].9   // VMCC W1 SPARE
        [43].10   // VMCC W1 SPARE
        [43].11   // VMCC W1 SPARE
        [60].14   // PANEL W3 JOG SPONGE ROLL FORWARD
        [43].14   // VMCC W1 SPARE
        [43].15   // VMCC W1 SPARE
        [56].0   // PANEL W2 BRUSH #1 AUTO Sw. Pos.
        [56].1   // PANEL W2 BRUSH #1 MANUAL Sw. Pos.
        [56].2   // PANEL W2 BRUSH #1 ON Sw. Pos.
        [56].3   // PANEL W2 BRUSH #1 OFF Sw. Pos.
        [62].15   // SPARE
        [62].10   // SPARE
        [62].12   // SPARE
        [56].8   // PANEL W2 SPONGE UNIT AUTO Sw. Pos.
        [56].9   // PANEL W2 SPONGE UNIT MANUAL Sw. Pos.
        [56].10   // PANEL W2 SPONGE UNIT ON Sw. Pos.
        [56].11   // PANEL W2 SPONGE UNIT OFF Sw. Pos.
        [56].12   // PANEL W2 AIR KNIFE AUTO Sw. Pos.
        [56].13   // PANEL W2 AIR KNIFE MANUAL Sw. Pos.
        [57].0   // PANEL W2 BRUSH #1 UPPER BRUSH CONVERGE Sw. Pos.
        [57].1   // PANEL W2 BRUSH #1 UPPER BRUSH RETRACT Sw. Pos.
        [58].8   // PANEL W2 AIR KNIFE BLOWER MODE OFF SS PANEL #W2
        [58].7   // PANEL W2 AIR KNIFE BLOWER MODE ON SS PANEL #W2
        [57].4   // PANEL W2 SPONGE UNIT UPPER SPONGE CONVERGE Sw. Pos.
        [57].5   // PANEL W2 SPONGE UNIT UPPER SPONGE RETRACT Sw. Pos.
        [57].6   // PANEL W2 BRUSH #1 LOWER BRUSH CONVERGE Sw. Pos.
        [57].7   // PANEL W2 BRUSH #1 LOWER BRUSH RETRACT Sw. Pos.
        [62].8   // PANEL W3 AIR KNIFE BLOWER MODE OFF SS PANEL #W3
        [62].7   // PANEL W3 AIR KNIFE BLOWER MODE ON SS PANEL #W3
        [57].10   // PANEL W2 SPONGE UNIT LOWER SPONGE CONVERGE Sw. Pos.
        [57].11   // PANEL W2 SPONGE UNIT LOWER SPONGE RETRACT Sw. Pos.
        [57].12   // PANEL W2 AIR KNIFE UNIT #1 CONVERGE Sw. Pos.
        [57].13   // PANEL W2 AIR KNIFE UNIT #1 RETRACT Sw. Pos.
        [57].14   // PANEL W2 AIR KNIFE UNIT #2 CONVERGE Sw. Pos.
        [57].15   // PANEL W2 AIR KNIFE UNIT #2 RETRACT Sw. Pos.
        [58].0   // PANEL W2 Cross break Reset Push-button
        [58].1   // PANEL W2 WATER SPRAYERS AUTO Sw. Pos.
        [58].2   // PANEL W2 WATER SPRAYERS MANUAL Sw. Pos.
        [58].3   // PANEL W2 WATER SPRAYERS ON Sw. Pos.
        [58].4   // PANEL W2 WATER SPRAYERS OFF Sw. Pos.
        [60].0   // PANEL W3 BRUSH #1 AUTO Sw. Pos.
        [60].1   // PANEL W3 BRUSH #1 MANUAL Sw. Pos.
        [60].2   // PANEL W3 BRUSH #1 ON Sw. Pos.
        [60].3   // PANEL W3 BRUSH #1 OFF Sw. Pos.
        [62].11   // SPARE